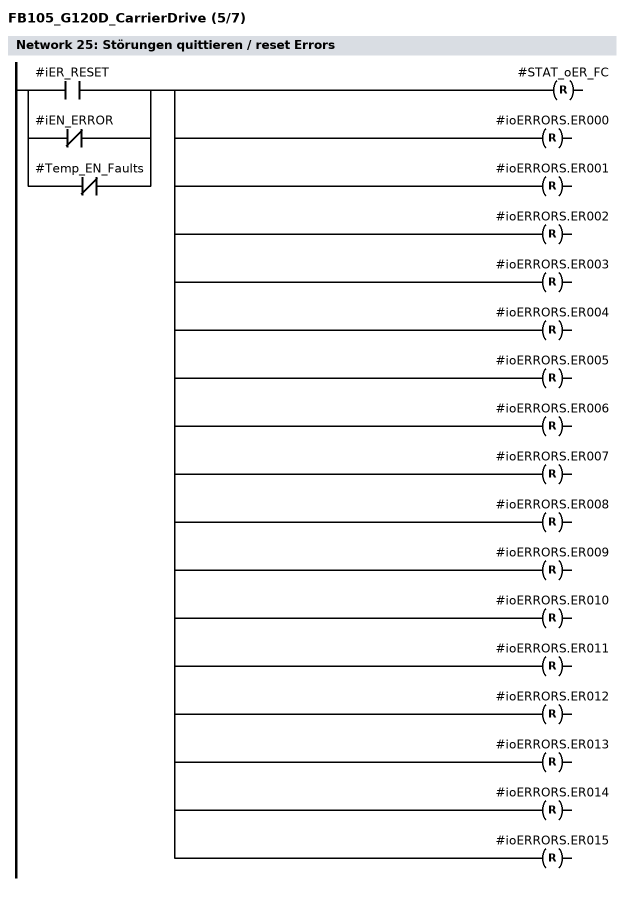
   RUNG wire#powerrail
      Contact( #iER_RESET )
      wire#w1
      R_Coil( #STAT_oER_FC )
   END_RUNG
   RUNG wire#powerrail
      I_Contact( #iEN_ERROR )
   END_RUNG wire#w1
   RUNG wire#powerrail
      I_Contact( #Temp_EN_Faults )
   END_RUNG wire#w1
   RUNG wire#w1
      R_Coil( #ioERRORS.ER000 )
   END_RUNG
   RUNG wire#w1
      R_Coil( #ioERRORS.ER001 )
   END_RUNG
   RUNG wire#w1
      R_Coil( #ioERRORS.ER002 )
   END_RUNG
   RUNG wire#w1
      R_Coil( #ioERRORS.ER003 )
   END_RUNG
   RUNG wire#w1
      R_Coil( #ioERRORS.ER004 )
   END_RUNG
   RUNG wire#w1
      R_Coil( #ioERRORS.ER005 )
   END_RUNG
   RUNG wire#w1
      R_Coil( #ioERRORS.ER006 )
   END_RUNG
   RUNG wire#w1
      R_Coil( #ioERRORS.ER007 )
   END_RUNG
   RUNG wire#w1
      R_Coil( #ioERRORS.ER008 )
   END_RUNG
   RUNG wire#w1
      R_Coil( #ioERRORS.ER009 )
   END_RUNG
   RUNG wire#w1
      R_Coil( #ioERRORS.ER010 )
   END_RUNG
   RUNG wire#w1
      R_Coil( #ioERRORS.ER011 )
   END_RUNG
   RUNG wire#w1
      R_Coil( #ioERRORS.ER012 )
   END_RUNG
   RUNG wire#w1
      R_Coil( #ioERRORS.ER013 )
   END_RUNG
   RUNG wire#w1
      R_Coil( #ioERRORS.ER014 )
   END_RUNG
   RUNG wire#w1
      R_Coil( #ioERRORS.ER015 )
   END_RUNG
   // the same network as SCL:
   IF #iER_RESET OR NOT #iEN_ERROR OR NOT #Temp_EN_Faults THEN
       #STAT_oER_FC := FALSE;
       #ioERRORS.ER000 := FALSE;
       #ioERRORS.ER001 := FALSE;
       #ioERRORS.ER002 := FALSE;
       #ioERRORS.ER003 := FALSE;
       #ioERRORS.ER004 := FALSE;
       #ioERRORS.ER005 := FALSE;
       #ioERRORS.ER006 := FALSE;
       #ioERRORS.ER007 := FALSE;
       #ioERRORS.ER008 := FALSE;
       #ioERRORS.ER009 := FALSE;
       #ioERRORS.ER010 := FALSE;
       #ioERRORS.ER011 := FALSE;
       #ioERRORS.ER012 := FALSE;
       #ioERRORS.ER013 := FALSE;
       #ioERRORS.ER014 := FALSE;
       #ioERRORS.ER015 := FALSE;
   END_IF;
END_REGION

REGION Network 26: Störungen / Errors
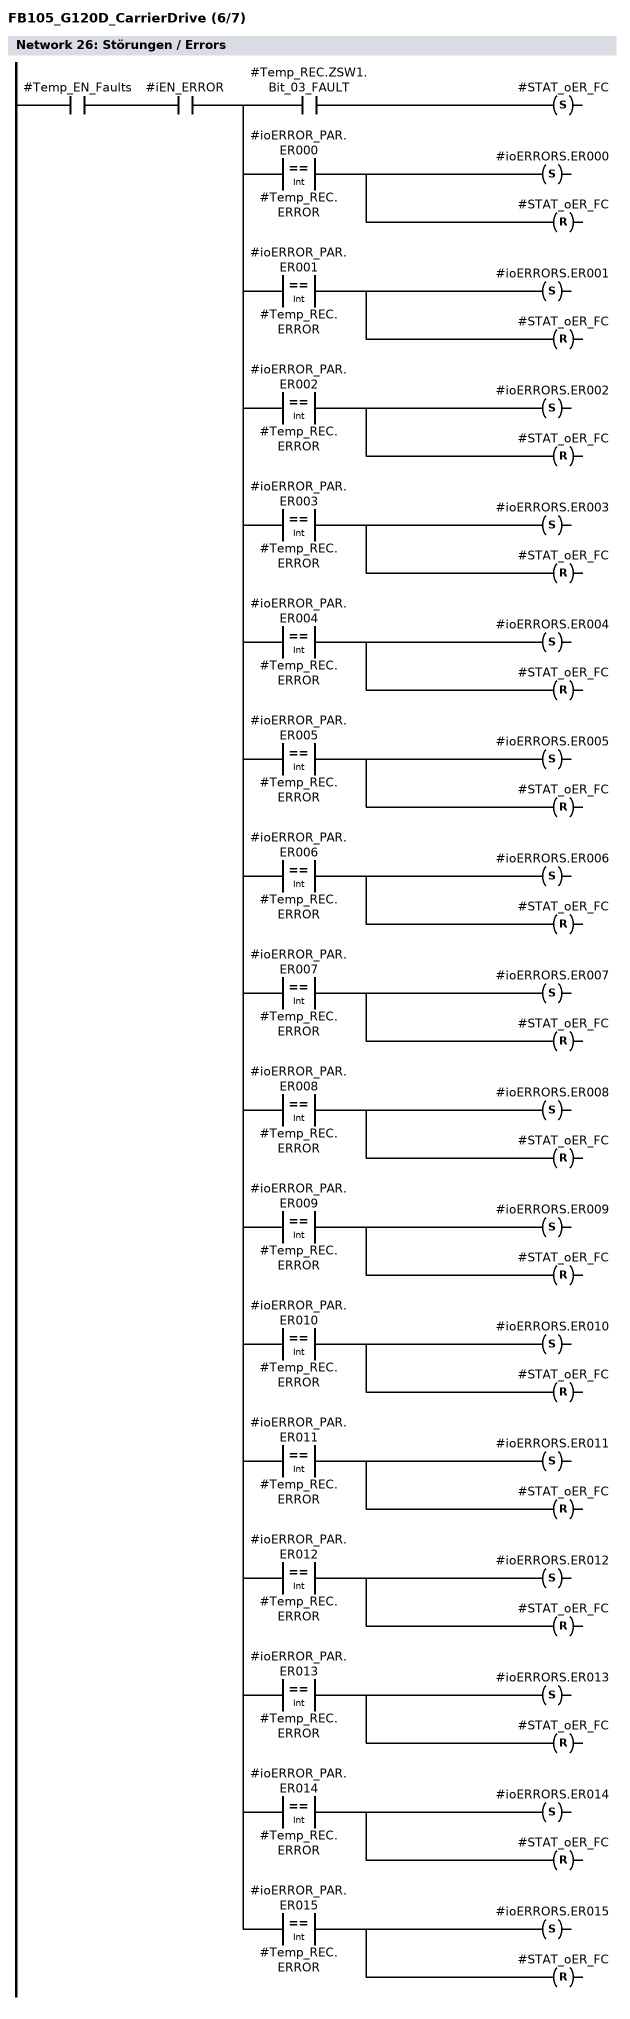
   RUNG wire#powerrail
      Contact( #Temp_EN_Faults )
      Contact( #iEN_ERROR )
      wire#w1
      Contact( #Temp_REC.ZSW1.Bit_03_FAULT )
      S_Coil( #STAT_oER_FC )
   END_RUNG
   RUNG wire#w1
      { S7_Templates := "SrcType := Int" } EQ_Contact(in1 := #ioERROR_PAR.ER000, in2 := #Temp_REC.ERROR)
      wire#w2
      S_Coil( #ioERRORS.ER000 )
   END_RUNG
   RUNG wire#w2
      R_Coil( #STAT_oER_FC )
   END_RUNG
   RUNG wire#w1
      { S7_Templates := "SrcType := Int" } EQ_Contact(in1 := #ioERROR_PAR.ER001, in2 := #Temp_REC.ERROR)
      wire#w3
      S_Coil( #ioERRORS.ER001 )
   END_RUNG
   RUNG wire#w3
      R_Coil( #STAT_oER_FC )
   END_RUNG
   RUNG wire#w1
      { S7_Templates := "SrcType := Int" } EQ_Contact(in1 := #ioERROR_PAR.ER002, in2 := #Temp_REC.ERROR)
      wire#w4
      S_Coil( #ioERRORS.ER002 )
   END_RUNG
   RUNG wire#w4
      R_Coil( #STAT_oER_FC )
   END_RUNG
   RUNG wire#w1
      { S7_Templates := "SrcType := Int" } EQ_Contact(in1 := #ioERROR_PAR.ER003, in2 := #Temp_REC.ERROR)
      wire#w5
      S_Coil( #ioERRORS.ER003 )
   END_RUNG
   RUNG wire#w5
      R_Coil( #STAT_oER_FC )
   END_RUNG
   RUNG wire#w1
      { S7_Templates := "SrcType := Int" } EQ_Contact(in1 := #ioERROR_PAR.ER004, in2 := #Temp_REC.ERROR)
      wire#w6
      S_Coil( #ioERRORS.ER004 )
   END_RUNG
   RUNG wire#w6
      R_Coil( #STAT_oER_FC )
   END_RUNG
   RUNG wire#w1
      { S7_Templates := "SrcType := Int" } EQ_Contact(in1 := #ioERROR_PAR.ER005, in2 := #Temp_REC.ERROR)
      wire#w7
      S_Coil( #ioERRORS.ER005 )
   END_RUNG
   RUNG wire#w7
      R_Coil( #STAT_oER_FC )
   END_RUNG
   RUNG wire#w1
      { S7_Templates := "SrcType := Int" } EQ_Contact(in1 := #ioERROR_PAR.ER006, in2 := #Temp_REC.ERROR)
      wire#w8
      S_Coil( #ioERRORS.ER006 )
   END_RUNG
   RUNG wire#w8
      R_Coil( #STAT_oER_FC )
   END_RUNG
   RUNG wire#w1
      { S7_Templates := "SrcType := Int" } EQ_Contact(in1 := #ioERROR_PAR.ER007, in2 := #Temp_REC.ERROR)
      wire#w9
      S_Coil( #ioERRORS.ER007 )
   END_RUNG
   RUNG wire#w9
      R_Coil( #STAT_oER_FC )
   END_RUNG
   RUNG wire#w1
      { S7_Templates := "SrcType := Int" } EQ_Contact(in1 := #ioERROR_PAR.ER008, in2 := #Temp_REC.ERROR)
      wire#w10
      S_Coil( #ioERRORS.ER008 )
   END_RUNG
   RUNG wire#w10
      R_Coil( #STAT_oER_FC )
   END_RUNG
   RUNG wire#w1
      { S7_Templates := "SrcType := Int" } EQ_Contact(in1 := #ioERROR_PAR.ER009, in2 := #Temp_REC.ERROR)
      wire#w11
      S_Coil( #ioERRORS.ER009 )
   END_RUNG
   RUNG wire#w11
      R_Coil( #STAT_oER_FC )
   END_RUNG
   RUNG wire#w1
      { S7_Templates := "SrcType := Int" } EQ_Contact(in1 := #ioERROR_PAR.ER010, in2 := #Temp_REC.ERROR)
      wire#w12
      S_Coil( #ioERRORS.ER010 )
   END_RUNG
   RUNG wire#w12
      R_Coil( #STAT_oER_FC )
   END_RUNG
   RUNG wire#w1
      { S7_Templates := "SrcType := Int" } EQ_Contact(in1 := #ioERROR_PAR.ER011, in2 := #Temp_REC.ERROR)
      wire#w13
      S_Coil( #ioERRORS.ER011 )
   END_RUNG
   RUNG wire#w13
      R_Coil( #STAT_oER_FC )
   END_RUNG
   RUNG wire#w1
      { S7_Templates := "SrcType := Int" } EQ_Contact(in1 := #ioERROR_PAR.ER012, in2 := #Temp_REC.ERROR)
      wire#w14
      S_Coil( #ioERRORS.ER012 )
   END_RUNG
   RUNG wire#w14
      R_Coil( #STAT_oER_FC )
   END_RUNG
   RUNG wire#w1
      { S7_Templates := "SrcType := Int" } EQ_Contact(in1 := #ioERROR_PAR.ER013, in2 := #Temp_REC.ERROR)
      wire#w15
      S_Coil( #ioERRORS.ER013 )
   END_RUNG
   RUNG wire#w15
      R_Coil( #STAT_oER_FC )
   END_RUNG
   RUNG wire#w1
      { S7_Templates := "SrcType := Int" } EQ_Contact(in1 := #ioERROR_PAR.ER014, in2 := #Temp_REC.ERROR)
      wire#w16
      S_Coil( #ioERRORS.ER014 )
   END_RUNG
   RUNG wire#w16
      R_Coil( #STAT_oER_FC )
   END_RUNG
   RUNG wire#w1
      { S7_Templates := "SrcType := Int" } EQ_Contact(in1 := #ioERROR_PAR.ER015, in2 := #Temp_REC.ERROR)
      wire#w17
      S_Coil( #ioERRORS.ER015 )
   END_RUNG
   RUNG wire#w17
      R_Coil( #STAT_oER_FC )
   END_RUNG
   // the same network as SCL:
   #_w1 := #Temp_EN_Faults AND #iEN_ERROR;
   IF #_w1 AND #Temp_REC.ZSW1.Bit_03_FAULT THEN #STAT_oER_FC := TRUE; END_IF;
   IF #_w1 AND (#ioERROR_PAR.ER000 = #Temp_REC.ERROR) THEN
       #ioERRORS.ER000 := TRUE;
       #STAT_oER_FC := FALSE;
   END_IF;
   IF #_w1 AND (#ioERROR_PAR.ER001 = #Temp_REC.ERROR) THEN
       #ioERRORS.ER001 := TRUE;
       #STAT_oER_FC := FALSE;
   END_IF;
   IF #_w1 AND (#ioERROR_PAR.ER002 = #Temp_REC.ERROR) THEN
       #ioERRORS.ER002 := TRUE;
       #STAT_oER_FC := FALSE;
   END_IF;
   IF #_w1 AND (#ioERROR_PAR.ER003 = #Temp_REC.ERROR) THEN
       #ioERRORS.ER003 := TRUE;
       #STAT_oER_FC := FALSE;
   END_IF;
   IF #_w1 AND (#ioERROR_PAR.ER004 = #Temp_REC.ERROR) THEN
       #ioERRORS.ER004 := TRUE;
       #STAT_oER_FC := FALSE;
   END_IF;
   IF #_w1 AND (#ioERROR_PAR.ER005 = #Temp_REC.ERROR) THEN
       #ioERRORS.ER005 := TRUE;
       #STAT_oER_FC := FALSE;
   END_IF;
   IF #_w1 AND (#ioERROR_PAR.ER006 = #Temp_REC.ERROR) THEN
       #ioERRORS.ER006 := TRUE;
       #STAT_oER_FC := FALSE;
   END_IF;
   IF #_w1 AND (#ioERROR_PAR.ER007 = #Temp_REC.ERROR) THEN
       #ioERRORS.ER007 := TRUE;
       #STAT_oER_FC := FALSE;
   END_IF;
   IF #_w1 AND (#ioERROR_PAR.ER008 = #Temp_REC.ERROR) THEN
       #ioERRORS.ER008 := TRUE;
       #STAT_oER_FC := FALSE;
   END_IF;
   IF #_w1 AND (#ioERROR_PAR.ER009 = #Temp_REC.ERROR) THEN
       #ioERRORS.ER009 := TRUE;
       #STAT_oER_FC := FALSE;
   END_IF;
   IF #_w1 AND (#ioERROR_PAR.ER010 = #Temp_REC.ERROR) THEN
       #ioERRORS.ER010 := TRUE;
       #STAT_oER_FC := FALSE;
   END_IF;
   IF #_w1 AND (#ioERROR_PAR.ER011 = #Temp_REC.ERROR) THEN
       #ioERRORS.ER011 := TRUE;
       #STAT_oER_FC := FALSE;
   END_IF;
   IF #_w1 AND (#ioERROR_PAR.ER012 = #Temp_REC.ERROR) THEN
       #ioERRORS.ER012 := TRUE;
       #STAT_oER_FC := FALSE;
   END_IF;
   IF #_w1 AND (#ioERROR_PAR.ER013 = #Temp_REC.ERROR) THEN
       #ioERRORS.ER013 := TRUE;
       #STAT_oER_FC := FALSE;
   END_IF;
   IF #_w1 AND (#ioERROR_PAR.ER014 = #Temp_REC.ERROR) THEN
       #ioERRORS.ER014 := TRUE;
       #STAT_oER_FC := FALSE;
   END_IF;
   IF #_w1 AND (#ioERROR_PAR.ER015 = #Temp_REC.ERROR) THEN
       #ioERRORS.ER015 := TRUE;
       #STAT_oER_FC := FALSE;
   END_IF;
END_REGION

REGION Network 27: OUT: Störung FU allgemein
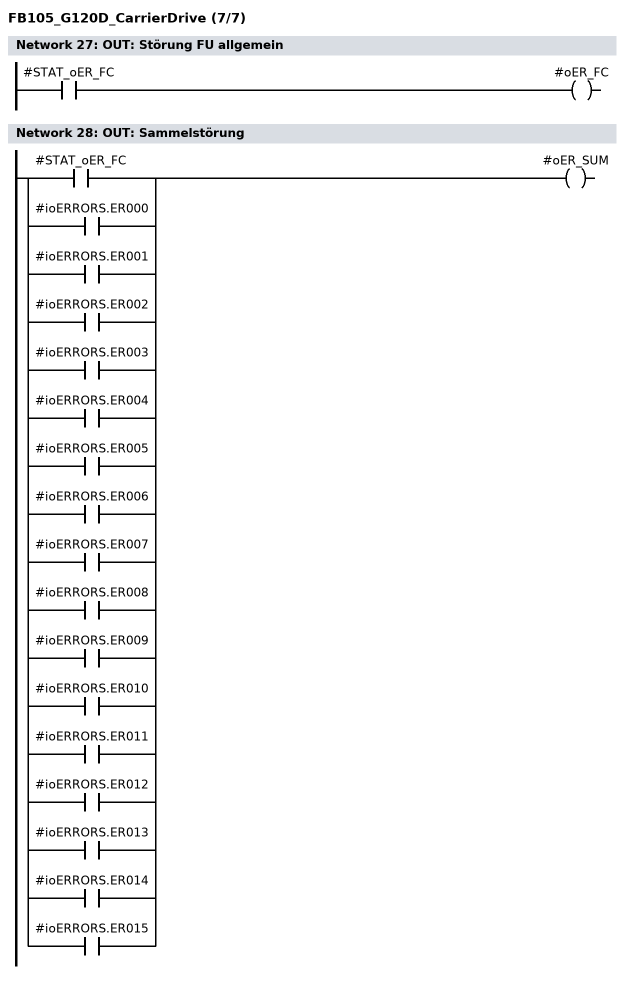
   RUNG wire#powerrail
      Contact( #STAT_oER_FC )
      Coil( #oER_FC )
   END_RUNG
   // the same network as SCL:
   #oER_FC := #STAT_oER_FC;
END_REGION

REGION Network 28: OUT: Sammelstörung
   RUNG wire#powerrail
      Contact( #STAT_oER_FC )
      wire#w1
      Coil( #oER_SUM )
   END_RUNG
   RUNG wire#powerrail
      Contact( #ioERRORS.ER000 )
   END_RUNG wire#w1
   RUNG wire#powerrail
      Contact( #ioERRORS.ER001 )
   END_RUNG wire#w1
   RUNG wire#powerrail
      Contact( #ioERRORS.ER002 )
   END_RUNG wire#w1
   RUNG wire#powerrail
      Contact( #ioERRORS.ER003 )
   END_RUNG wire#w1
   RUNG wire#powerrail
      Contact( #ioERRORS.ER004 )
   END_RUNG wire#w1
   RUNG wire#powerrail
      Contact( #ioERRORS.ER005 )
   END_RUNG wire#w1
   RUNG wire#powerrail
      Contact( #ioERRORS.ER006 )
   END_RUNG wire#w1
   RUNG wire#powerrail
      Contact( #ioERRORS.ER007 )
   END_RUNG wire#w1
   RUNG wire#powerrail
      Contact( #ioERRORS.ER008 )
   END_RUNG wire#w1
   RUNG wire#powerrail
      Contact( #ioERRORS.ER009 )
   END_RUNG wire#w1
   RUNG wire#powerrail
      Contact( #ioERRORS.ER010 )
   END_RUNG wire#w1
   RUNG wire#powerrail
      Contact( #ioERRORS.ER011 )
   END_RUNG wire#w1
   RUNG wire#powerrail
      Contact( #ioERRORS.ER012 )
   END_RUNG wire#w1
   RUNG wire#powerrail
      Contact( #ioERRORS.ER013 )
   END_RUNG wire#w1
   RUNG wire#powerrail
      Contact( #ioERRORS.ER014 )
   END_RUNG wire#w1
   RUNG wire#powerrail
      Contact( #ioERRORS.ER015 )
   END_RUNG wire#w1
   // the same network as SCL:
   #oER_SUM := #STAT_oER_FC OR #ioERRORS.ER000 OR #ioERRORS.ER001 OR #ioERRORS.ER002 OR #ioERRORS.ER003 OR #ioERRORS.ER004 OR #ioERRORS.ER005 OR #ioERRORS.ER006 OR #ioERRORS.ER007 OR #ioERRORS.ER008 OR #ioERRORS.ER009 OR #ioERRORS.ER010 OR #ioERRORS.ER011 OR #ioERRORS.ER012 OR #ioERRORS.ER013 OR #ioERRORS.ER014 OR #ioERRORS.ER015;
END_REGION

REGION Network 29: ENDE / END
   // ################################ ENDE ############################### / ###################################### END #####################################
END_REGION
END_FUNCTION_BLOCK

FUNCTION_BLOCK "FB1110_Red_Green_LED"   // FB1110, LAD
{ S7_Optimized_Access := 'TRUE' }
VERSION : 0.1
   VAR_INPUT
      Red : Bool;
      Green : Bool;
   END_VAR
   VAR
      instWRREC : WRREC;
      statWRREC_LEDByte : Byte;
   END_VAR
BEGIN

REGION Network 1: Red LED
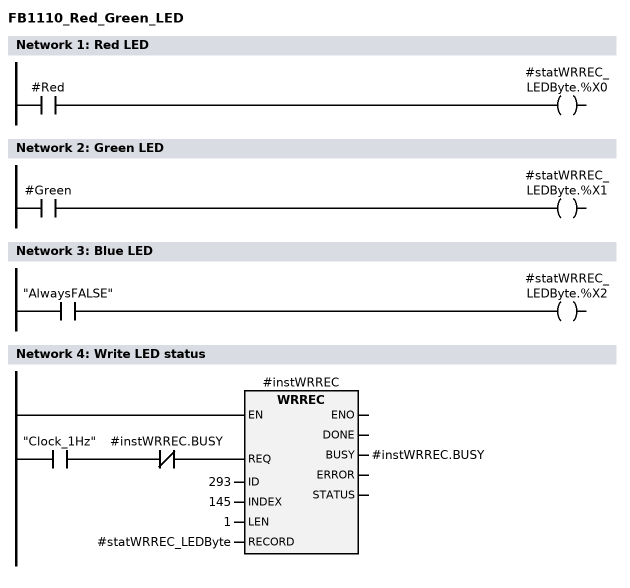
   RUNG wire#powerrail
      Contact( #Red )
      Coil( #statWRREC_LEDByte.%X0 )
   END_RUNG
   // the same network as SCL:
   #statWRREC_LEDByte.%X0 := #Red;
END_REGION

REGION Network 2: Green LED
   RUNG wire#powerrail
      Contact( #Green )
      Coil( #statWRREC_LEDByte.%X1 )
   END_RUNG
   // the same network as SCL:
   #statWRREC_LEDByte.%X1 := #Green;
END_REGION

REGION Network 3: Blue LED
   RUNG wire#powerrail
      Contact( "AlwaysFALSE" )
      Coil( #statWRREC_LEDByte.%X2 )
   END_RUNG
   // the same network as SCL:
   #statWRREC_LEDByte.%X2 := "AlwaysFALSE";
END_REGION

REGION Network 4: Write LED status
   #instWRREC(REQ := "Clock_1Hz" AND NOT #instWRREC.BUSY,   // WRREC
              ID := 293,
              INDEX := 145,
              LEN := 1,
              RECORD := #statWRREC_LEDByte,
              BUSY => #instWRREC.BUSY);
END_REGION

REGION Network 5: End
END_REGION
END_FUNCTION_BLOCK

// folder: 03_FB'S/DIAGNOSTICS

FUNCTION_BLOCK "FB1000_Default_SupervisionFB"   // FB1000, ProDiag
{ S7_Optimized_Access := 'TRUE' }
   VAR
      State : SV_FB_State;
   END_VAR
   VAR_TEMP
      t_TempSvStateUDT : SV_State;
      t_TempAlarmInstance : <type 200004f>;
      t_TempAsocValue1 : Variant;
      t_TempAsocValue2 : Variant;
      t_TempAsocValue3 : Variant;
   END_VAR
BEGIN
END_FUNCTION_BLOCK

FUNCTION_BLOCK "FB1001_EMS_BreakerStatus"   // FB1001, LAD
TITLE = Monitoring Fuse
{ S7_Optimized_Access := 'TRUE' }
AUTHOR : Siemens
FAMILY : LSimoveC
VERSION : 1.0
// © 2018 Siemens AG 
// SIMOVE Carrier Control
   VAR_INPUT
      Diag : Variant;   // Diagnosis signal of the selectivity module
   END_VAR
   VAR_OUTPUT
      Channel1 : Bool;   // Channel 1 active
      Channel2 : Bool;   // Channel 2 active
      Channel3 : Bool;   // Channel 3 active
      Channel4 : Bool;   // Channel 4 active
      CollectiveError : Bool;   // Collective error of the selectivity module
   END_VAR
   VAR
      instDiagBreaker : "FB1002_LSimoveC_DiagBreaker";
      instTimeout : TON_TIME;
      statError : Bool;
   END_VAR
   VAR_TEMP
      tempDone : Bool;
      tempBusy : Bool;
      tempChannelState : Byte;
      tempStatus : Word;
      tempDiag : Bool;
      tempInt : Int;
      tempModuleOK : Bool;
      tempHW : Hw_Any;
      tempDiagInfo : DIS;
      tempUInt : UInt;
      tempTimeout : Bool;
   END_VAR
BEGIN

REGION Network 1: Change journal
   // =============================================================================
   // Siemens AG
   // (c)Copyright 2018 Alle Rechte vorbehalten
   // -----------------------------------------------------------------------------
   // Bibliothek: LSimoveC
   // Funktion: Der FB wertet den Status-Ausgang eines SITOP-Selektivitätsmoduls aus. Der Status-Ausgang liefert ein Signal, das den Zustand der Verbaucherkreise seriell codiert. Der Baustein decodiert das Signal und stellt den Status der Verbraucherkreise als Einzelsignale zur Verfügung.
   // -----------------------------------------------------------------------------
   // Änderungsjournal:
   // V1.0  01.02.2018  Neuerstellung
   // =============================================================================
END_REGION

REGION Network 2: Determine block error
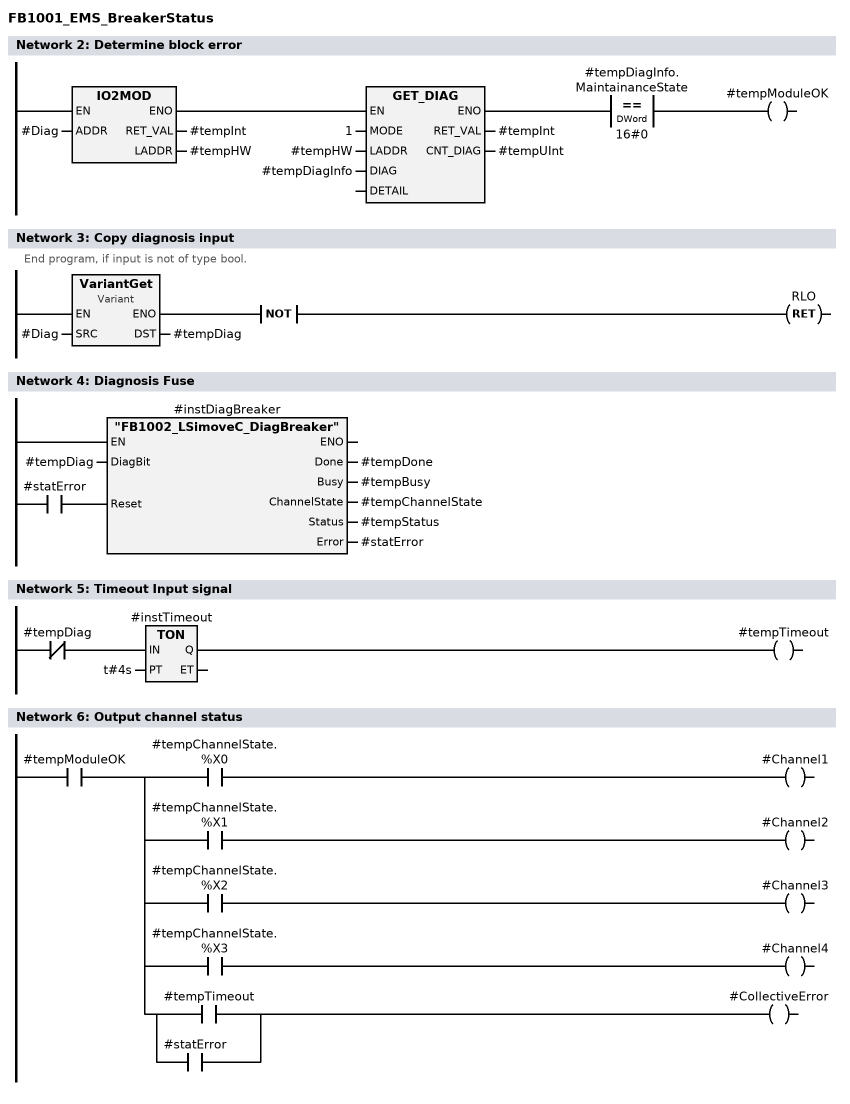
   // ENO of a box is taken as its EN; it also drops when the box reports an error
   #tempInt := IO2MOD(ADDR := #Diag, LADDR => #tempHW);
   #tempInt := GET_DIAG(MODE := 1, LADDR := #tempHW, DIAG := #tempDiagInfo, CNT_DIAG => #tempUInt);
   #tempModuleOK := #tempDiagInfo.MaintainanceState = 16#0;
END_REGION

REGION Network 3: Copy diagnosis input
   // End program, if input is not of type bool.
   // no SCL statement known for VariantGet: written as a call
   // ENO of a box is taken as its EN; it also drops when the box reports an error
   VariantGet(src := #Diag, dst => #tempDiag);
   IF NOT TRUE THEN
       ENO := TRUE;
       RETURN;
   END_IF;
END_REGION

REGION Network 4: Diagnosis Fuse
   RUNG wire#powerrail
      #instDiagBreaker(Reset := wire#w1, DiagBit := #tempDiag, Done => #tempDone, Busy => #tempBusy, ChannelState => #tempChannelState, Status => #tempStatus, Error => #statError)
   END_RUNG
   RUNG wire#powerrail
      Contact( #statError )
   END_RUNG wire#w1
   // the same network as SCL:
   #instDiagBreaker(DiagBit := #tempDiag,   // "FB1002_LSimoveC_DiagBreaker"
                    Reset := #statError,
                    Done => #tempDone,
                    Busy => #tempBusy,
                    ChannelState => #tempChannelState,
                    Status => #tempStatus,
                    Error => #statError);
END_REGION

REGION Network 5: Timeout Input signal
   #instTimeout(IN := NOT #tempDiag, PT := t#4s);   // TON
   #tempTimeout := #instTimeout.Q;
END_REGION

REGION Network 6: Output channel status
   RUNG wire#powerrail
      Contact( #tempModuleOK )
      wire#w1
      Contact( #tempChannelState.%X0 )
      Coil( #Channel1 )
   END_RUNG
   RUNG wire#w1
      Contact( #tempChannelState.%X1 )
      Coil( #Channel2 )
   END_RUNG
   RUNG wire#w1
      Contact( #tempChannelState.%X2 )
      Coil( #Channel3 )
   END_RUNG
   RUNG wire#w1
      Contact( #tempChannelState.%X3 )
      Coil( #Channel4 )
   END_RUNG
   RUNG wire#w1
      Contact( #tempTimeout )
      wire#w2
      Coil( #CollectiveError )
   END_RUNG
   RUNG wire#w1
      Contact( #statError )
   END_RUNG wire#w2
   // the same network as SCL:
   #Channel1 := #tempModuleOK AND #tempChannelState.%X0;
   #Channel2 := #tempModuleOK AND #tempChannelState.%X1;
   #Channel3 := #tempModuleOK AND #tempChannelState.%X2;
   #Channel4 := #tempModuleOK AND #tempChannelState.%X3;
   #CollectiveError := #tempModuleOK AND (#tempTimeout OR #statError);
END_REGION
END_FUNCTION_BLOCK

FUNCTION_BLOCK "FB1002_LSimoveC_DiagBreaker"   // FB1002, SCL
TITLE = DiagnoseSicherung
{ S7_Optimized_Access := 'FALSE' }
AUTHOR : Siemens
FAMILY : LSimoveC
VERSION : 2.3
// © 2018 Siemens AG 
// SIMOVE Carrier Control
   VAR_INPUT
      DiagBit : Bool;   // Input through which the signal of the status output of the selectivity module is read
      Reset : Bool;   // A positive edge triggers a reset. All parameters are reset.
   END_VAR
   VAR_OUTPUT
      Done : Bool;   // Done = 1: A telegram was evaluated completely and without errors. Done = 0: telegram evaluation is running or no signal is detected at the input "impulse".
      Busy : Bool;   // Busy = 1: Function module "LSitop_PseDiag" is active. Busy = 0: if done=1, a telegram was evaluated completely and without error.
      ChannelState : Byte;   // State of the outputs 1 to 4.
      Status : Word;   // Status display: if error=1, the error number for one cycle is displayed at the output "status". if error=0, the value 16 # 0000 is displayed at the output "status".
      Error : Bool;   // Error=1: an error has occured during the execution of the routine. The value error=1 is set for one cycle. if error=0: no error.
   END_VAR
   VAR
      statImpulseOld : Bool;
      statResetOld : Bool;
      statTimeSaver : Struct
         TimeTckRisingEdge : Time;
         TimeTckFallingEdge : Time;
         RisingEdgeDetected : Bool;
         FallingEdgeDetected : Bool;
         stateEdge : Int := 0;
      END_STRUCT;
      statDeltaTimeImpulse : Time;
      statDeltaTimePause : Time;
      statStartImpulseDetected : Bool;
      statImpulseDetected : Bool;
      statChannelState : Byte;
      statTimePauseSave0 : Time;
      statTimePauseSave1 : Time;
      statTimePauseSave2 : Time;
      statTimePauseSave3 : Time;
      statTimePauseSave4 : Time;
      statTimeImpulseSave0 : Time;
      statTimeImpulseSave1 : Time;
      statTimeImpulseSave2 : Time;
      statTimeImpulseSave3 : Time;
      statTimeImpulseSave4 : Time;
      statFrameImulseDetected : Bool;
      statNumberOfImpulses : Int;
      statChannelActive1 : Bool;
      statChannelActive2 : Bool;
      statChannelActive3 : Bool;
      statChannelActive4 : Bool;
      statCountChannelPos : Int;
      statCurrentPos1 : Int;
      statCurrentPos2 : Int;
      statCurrentPos3 : Int;
      statCurrentPos4 : Int;
      statTimeToImpulse : Time;
      statTimePause : Time;
      statTimeImpulse : Time;
      statTimeFrame : Time;
      statFrameOk : Bool;
      statCycleTimeNok : Bool;
      statSysTime : Time;
      statSysTimeOld : Time;
      statDeltaSysTime : Time;
      instSysTimer : TON_TIME;
      statSysTimerStart : Bool;
      statSysTimerStop : Bool;
      statStatus : Word;
      statIndex : Int;
      statSysTimerRun : Time;
      instWatchDogTimerRising : TON_TIME;
      statWatchDogTimerRisingStart : Bool;
      statWatchDogTimerRisingStop : Bool;
      statWatchDogTimerRisingRun : Time;
      statResetRequest : Bool;
      instWatchDogTimerFalling : TON_TIME;
      statWatchDogTimerFallingStart : Bool;
      statWatchDogTimerFallingStop : Bool;
      statWatchDogTimerFallingRun : Time;
   END_VAR
   VAR_TEMP
      tempLatchTime : Time;
   END_VAR
   VAR CONSTANT
      STATE_IDLE : Int := 0;
      STATE_EVALUATION : Int := 1;
      STATE_ERROR : Int := 2;
      TIME_FRAME_MAX : Time := T#2850ms;
      TIME_FRAME_MIN : Time := T#2650ms;
      TIME_STARTIMPULSE_MAX : Time := T#600ms;
      TIME_STARTIMPULSE_MIN : Time := T#400ms;
      TIME_IMPULSE_MIN : Time := T#150ms;
      TIME_IMPULSE_MAX : Time := T#350ms;
      TIME_PAUSE1_MIN : Time := T#150ms;
      TIME_PAUSE1_MAX : Time := T#350ms;
      TIME_PAUSE2_MIN : Time := T#650ms;
      TIME_PAUSE2_MAX : Time := T#850ms;
      TIME_PAUSE3_MIN : Time := T#1150ms;
      TIME_PAUSE3_MAX : Time := T#1350ms;
      TIME_PAUSE4_MIN : Time := T#1650ms;
      TIME_PAUSE4_MAX : Time := T#1850ms;
      TIME_PAUSE_FRAME_MAX : Time := T#2350ms;
      TIME_PAUSE_FRAME_MIN : Time := T#2150ms;
      TIME_CONST_0 : Time := T#0ms;
      TIME_CONST_102 : Time := T#102ms;
      CONST_STATE_RISING_EDGE : Int := 15;
      CONST_STATE_FALLING_EDGE : Int := 16;
      CONST_WORD_0 : Word := 16#0000;
      CONST_BYTE_0 : Byte := 16#00;
      CONST_INT_0 : Int := 0;
      CONST_CHANNEL_POS4 : Int := 4;
      CONST_CHANNEL_POS1 : Int := 1;
      CONST_CHANNEL_POS2 : Int := 2;
      CONST_CHANNEL_POS3 : Int := 3;
      CONST_WATCHDOG_TIMER : Time := T#6s;
      CONST_CYCLETIME_TIMER : Time := t#4s;
      CONST_ERROR_CYCLETIME_TIMER : Word := 16#8001;
      CONST_ERROR_WATCHDOG_TIMER : Word := 16#8002;
   END_VAR
BEGIN
   //=============================================================================
   //SIEMENES AG
   //(c)Copyright 2017 All Rights Reserved
   //-----------------------------------------------------------------------------
   //Library:       LSitop
   //Tested with:   (S7-1500)
   //Engineering:    TIA Portal V14
   //Restrictions:   call in cyclic main OB
   //Requirements:
   //Functionality: evaluates the signal of status output (S) of SITOP PSE200U 
   //               ....
   //
   //-----------------------------------------------------------------------------
   //Change log table:
   //Version  Date       Expert in charge Changes applied
   //02.03.01 24.05.2017 (DF CS SD CCC OS) Third released version
   //=============================================================================

   // Calculate cycle time
   #statSysTime:=TIME_TCK();
   #statDeltaSysTime := #statSysTime - #statSysTimeOld;

   IF (#statDeltaSysTime < t#0ms)
   THEN
       #statDeltaSysTime := #statDeltaSysTime + T#2147483647ms;

       IF (#statDeltaSysTime < #TIME_CONST_0)
       THEN
           #statCycleTimeNok := true;
           #statSysTimeOld := #statSysTime;
           RETURN;
       ELSE
           #statCycleTimeNok := false;
       END_IF;

   ELSIF (#statDeltaSysTime >= #TIME_CONST_102)
   THEN
       #statCycleTimeNok := true;
       #statSysTimerStart := true;
   ELSE
       #statCycleTimeNok := false;
       #statSysTimerStart := false;
   END_IF;

   //Rising edge at reset input

   IF ((#Reset = true)
       AND (#statResetOld = false))
   THEN
       #statSysTimerStart := false;
       #statWatchDogTimerRisingStart := false;
       #statWatchDogTimerFallingStart := false;
       #statResetRequest := true;
       #statIndex := #STATE_IDLE;
   END_IF;

   //Rising edge at impulse input
   IF ((#DiagBit = True)
       AND (#statImpulseOld = False))
   THEN
       #tempLatchTime := TIME_TCK();
       #statTimeSaver.RisingEdgeDetected := true;
       #statTimeSaver.stateEdge := #CONST_STATE_RISING_EDGE;
       #statTimeSaver.TimeTckRisingEdge := #tempLatchTime;
       #statWatchDogTimerRisingStart := true;
       #statWatchDogTimerFallingStart := false;

       IF (#Busy = false)
       THEN
           #Busy := true;
           #Done := false;
           #Error := false;
           #Status := #CONST_WORD_0;
       END_IF;

       IF ((#statCycleTimeNok = false)
           AND (#statResetRequest = false))
       THEN
           #statIndex := #STATE_EVALUATION;
       END_IF;

   END_IF;

   //Falling edge at impulse input
   IF ((#DiagBit = False)
       AND (#statImpulseOld = True))
   THEN
       #tempLatchTime := TIME_TCK();
       #statTimeSaver.FallingEdgeDetected := true;
       #statTimeSaver.stateEdge := #CONST_STATE_FALLING_EDGE;
       #statTimeSaver.TimeTckFallingEdge := #tempLatchTime;

       #statWatchDogTimerFallingStart := true;
       #statWatchDogTimerRisingStart := false;

       IF ((#statCycleTimeNok = FALSE)
           AND (#statResetRequest = false))
       THEN
           #statIndex := #STATE_EVALUATION;
       END_IF;

   END_IF;

   IF ((#statTimeSaver.FallingEdgeDetected = false)
       AND (#statTimeSaver.RisingEdgeDetected = FALSE))
   THEN
       #statWatchDogTimerRisingStart := true;
       #statWatchDogTimerFallingStart := true;
   END_IF;

   CASE #statIndex OF
       #STATE_IDLE:  // IDLE_STATE
           #Done := false;
           #Error := false;
           #Busy := false;
           #Status := #CONST_WORD_0;
           #statStatus := #CONST_WORD_0;
           #ChannelState := #CONST_BYTE_0;
           #statChannelState := #CONST_BYTE_0;
           #statFrameOk := false;
           #statCycleTimeNok := false;
           #statStartImpulseDetected := false;
           #statFrameImulseDetected := false;
           #statResetRequest := false;
           #statTimeSaver.FallingEdgeDetected := false;
           #statTimeSaver.RisingEdgeDetected := false;

       #STATE_EVALUATION:  //State: impulse detection

           //Delta time calculation
           IF ((#statTimeSaver.RisingEdgeDetected = True)
               AND (#statTimeSaver.FallingEdgeDetected = True))
           THEN

               IF (#statTimeSaver.stateEdge = #CONST_STATE_RISING_EDGE) //pos. edge, evaluate delta pause
               THEN
                   #statDeltaTimePause := #statTimeSaver.TimeTckRisingEdge - #statTimeSaver.TimeTckFallingEdge;

                   IF (#statDeltaTimePause < #TIME_CONST_0)
                   THEN
                       #statDeltaTimePause := #statDeltaTimePause + T#2147483647ms;

                       IF (#statDeltaTimePause < #TIME_CONST_0)
                       THEN
                           #statIndex := #STATE_IDLE;
                           #statTimeSaver.FallingEdgeDetected := false;
                           RETURN;
                       END_IF;

                   ELSIF (#statDeltaTimePause > #TIME_FRAME_MAX)
                   THEN
                       #statIndex := #STATE_IDLE;
                       #statTimeSaver.FallingEdgeDetected := false;
                       RETURN;
                   END_IF;
                   #statTimeSaver.FallingEdgeDetected := false;
               END_IF;

               IF (#statTimeSaver.stateEdge = #CONST_STATE_FALLING_EDGE) // neg. edge, evaluate delta impulse
               THEN
                   #statImpulseDetected := true;
                   #statDeltaTimeImpulse := #statTimeSaver.TimeTckFallingEdge - #statTimeSaver.TimeTckRisingEdge;

                   IF (#statDeltaTimeImpulse < #TIME_CONST_0)
                   THEN
                       #statDeltaTimeImpulse := #statDeltaTimeImpulse + T#2147483647ms;

                       IF (#statDeltaTimeImpulse < #TIME_CONST_0)
                       THEN
                           #statIndex := #STATE_IDLE;
                           #statTimeSaver.RisingEdgeDetected := false;
                           RETURN;
                       END_IF;

                   ELSIF (#statDeltaTimeImpulse > #TIME_FRAME_MAX)
                   THEN
                       #statIndex := #STATE_IDLE;
                       #statTimeSaver.RisingEdgeDetected := false;
                       RETURN;
                   END_IF;
                   #statTimeSaver.RisingEdgeDetected := false;
               END_IF;
           END_IF;

           //Start bit detection
           IF ((#statDeltaTimeImpulse >= #TIME_STARTIMPULSE_MIN)
               AND (#statDeltaTimeImpulse <= #TIME_STARTIMPULSE_MAX))
               AND (#statImpulseDetected = True)
           THEN
               #statImpulseDetected := False;
               #statNumberOfImpulses := #CONST_INT_0;
               #statCountChannelPos := #CONST_INT_0;

               IF (#statCurrentPos1 = #CONST_INT_0)
               THEN
                   #statTimeImpulseSave1 := #TIME_CONST_0;
                   #statTimePauseSave1 := #TIME_CONST_0;
               END_IF;

               IF (#statCurrentPos2 = #CONST_INT_0)
               THEN
                   #statTimeImpulseSave2 := #TIME_CONST_0;
                   #statTimePauseSave2 := #TIME_CONST_0;
               END_IF;

               IF (#statCurrentPos3 = #CONST_INT_0)
               THEN
                   #statTimeImpulseSave3 := #TIME_CONST_0;
                   #statTimePauseSave3 := #TIME_CONST_0;
               END_IF;

               IF (#statCurrentPos4 = #CONST_INT_0)
               THEN
                   #statTimeImpulseSave4 := #TIME_CONST_0;
                   #statTimePauseSave4 := #TIME_CONST_0;
               END_IF;

               #statTimePauseSave0 := #statDeltaTimePause;
               #statTimeImpulseSave0 := #statDeltaTimeImpulse;

               // get time in sum of imulses
               #statTimeImpulse := #statTimeImpulseSave0 + #statTimeImpulseSave1 + #statTimeImpulseSave2 + #statTimeImpulseSave3 + #statTimeImpulseSave4;

               //get time in sum of pauses
               #statTimePause := #statTimePauseSave0 + #statTimePauseSave1 + #statTimePauseSave2 + #statTimePauseSave3 + #statTimePauseSave4;

               // get length of frame
               #statTimeFrame := #statTimeImpulse + #statTimePause;

               IF ((#statTimeFrame >= #TIME_FRAME_MIN)
                   AND (#statTimeFrame <= #TIME_FRAME_MAX)
                   AND (#statTimeToImpulse <= #TIME_FRAME_MAX))
               THEN
                   #statFrameOk := true;
               END_IF;

               IF ((#statFrameOk = TRUE)
                   AND (#statCycleTimeNok = FALSE))
               THEN
                   // take over data
                   #Done := true;
                   #Busy := false;
                   #statFrameOk := false;

                   IF (#statChannelActive1 = true)
                   THEN
                       #statChannelState.%X0 := false;
                   ELSE
                       #statChannelState.%X0 := true;
                   END_IF;

                   IF (#statChannelActive2 = true)
                   THEN
                       #statChannelState.%X1 := false;
                   ELSE
                       #statChannelState.%X1 := true;
                   END_IF;

                   IF (#statChannelActive3 = true)
                   THEN
                       #statChannelState.%X2 := false;
                   ELSE
                       #statChannelState.%X2 := true;
                   END_IF;

                   IF (#statChannelActive4 = true)
                   THEN
                       #statChannelState.%X3 := false;
                   ELSE
                       #statChannelState.%X3 := true;
                   END_IF;

                   #ChannelState := #statChannelState;
               END_IF;


               // channel 4 ok
               IF ((#statDeltaTimePause >= #TIME_PAUSE1_MIN)
                   AND (#statDeltaTimePause <= #TIME_PAUSE1_MAX))
               THEN
                   #statChannelActive4 := true;
                   // channel 4 ok not ok
               ELSIF ((#statDeltaTimePause >= #TIME_PAUSE2_MIN)
                   AND (#statDeltaTimePause <= #TIME_PAUSE2_MAX))
               THEN
                   #statChannelActive4 := false;
                   // channel 3 and 4 not ok    
               ELSIF ((#statDeltaTimePause >= #TIME_PAUSE3_MIN)
                   AND (#statDeltaTimePause <= #TIME_PAUSE3_MAX))
               THEN
                   #statChannelActive3 := false;
                   #statChannelActive4 := false;
                   // channel 2, 3, 4 not ok
               ELSIF ((#statDeltaTimePause >= #TIME_PAUSE4_MIN)
                   AND (#statDeltaTimePause <= #TIME_PAUSE4_MAX))
               THEN
                   #statChannelActive2 := false;
                   #statChannelActive3 := false;
                   #statChannelActive4 := false;
                   // channel 1, 2, 3, 4 not ok
               ELSIF ((#statDeltaTimePause >= #TIME_PAUSE_FRAME_MIN)
                   AND (#statDeltaTimePause <= #TIME_PAUSE_FRAME_MAX))
               THEN
                   #statChannelActive1 := false;
                   #statChannelActive2 := false;
                   #statChannelActive3 := false;
                   #statChannelActive4 := false;
               END_IF;

               #statCountChannelPos := #CONST_CHANNEL_POS4;

               #statCurrentPos1 := #CONST_INT_0;
               #statCurrentPos2 := #CONST_INT_0;
               #statCurrentPos3 := #CONST_INT_0;
               #statCurrentPos4 := #CONST_INT_0;

           // Imulse bit detection
           ELSIF ((#statDeltaTimeImpulse >= #TIME_IMPULSE_MIN)
               AND (#statDeltaTimeImpulse <= #TIME_IMPULSE_MAX))
               AND (#statImpulseDetected = True)
           THEN
               #statImpulseDetected := False;
               #statFrameImulseDetected := true;
           END_IF;

           //Channel detection
           IF #statFrameImulseDetected = TRUE
           THEN
               #statFrameImulseDetected := FALSE;

               IF (#statCountChannelPos = #CONST_CHANNEL_POS4)
               THEN
                   #statCurrentPos1 := #statCountChannelPos;
                   #statTimeImpulseSave1 := #statDeltaTimeImpulse;
                   #statTimePauseSave1 := #statDeltaTimePause;
                   #statTimeToImpulse := #TIME_CONST_0;
                   #statTimeToImpulse := #statTimeToImpulse + #statDeltaTimeImpulse + #statDeltaTimePause;

                   //channel 1 ok
                   IF ((#statDeltaTimePause >= #TIME_PAUSE1_MIN)
                       AND (#statDeltaTimePause <= #TIME_PAUSE1_MAX))
                   THEN
                       #statChannelActive1 := true;
                       #statCountChannelPos := #CONST_CHANNEL_POS1; // Pos 1 detected
                   END_IF;

                   // channel 1 not ok
                   IF ((#statDeltaTimePause >= #TIME_PAUSE2_MIN)
                       AND (#statDeltaTimePause <= #TIME_PAUSE2_MAX))
                   THEN
                       #statChannelActive1 := false;
                       #statChannelActive2 := true;
                       #statCountChannelPos := #CONST_CHANNEL_POS2; // go to next Pos 2
                   END_IF;

                   // channel 1 and 2 not ok
                   IF ((#statDeltaTimePause >= #TIME_PAUSE3_MIN)
                       AND (#statDeltaTimePause <= #TIME_PAUSE3_MAX))
                   THEN
                       #statChannelActive1 := false;
                       #statChannelActive2 := false;
                       #statChannelActive3 := true;
                       #statCountChannelPos := #CONST_CHANNEL_POS2; // go to next Pos 2
                   END_IF;

                   // channel 1, 2 and 3 not ok
                   IF ((#statDeltaTimePause >= #TIME_PAUSE4_MIN)
                       AND (#statDeltaTimePause <= #TIME_PAUSE4_MAX))
                   THEN
                       #statChannelActive1 := false;
                       #statChannelActive2 := false;
                       #statChannelActive3 := FALSE;
                       #statChannelActive4 := true;
                       #statCountChannelPos := #CONST_INT_0;
                   END_IF;

               ELSIF (#statCountChannelPos = #CONST_CHANNEL_POS1)
               THEN
                   #statCurrentPos2 := #statCountChannelPos;
                   #statTimeImpulseSave2 := #statDeltaTimeImpulse;
                   #statTimePauseSave2 := #statDeltaTimePause;
                   #statTimeToImpulse := #statTimeToImpulse + #statDeltaTimeImpulse + #statDeltaTimePause;

                   IF ((#statDeltaTimePause >= #TIME_PAUSE1_MIN)
                       AND (#statDeltaTimePause <= #TIME_PAUSE1_MAX))
                   THEN
                       #statChannelActive2 := true;
                       #statCountChannelPos := #CONST_CHANNEL_POS2; // go to next pos 2
                   END_IF;

                   IF ((#statDeltaTimePause >= #TIME_PAUSE2_MIN)
                       AND (#statDeltaTimePause <= #TIME_PAUSE2_MAX))
                   THEN
                       #statChannelActive2 := false;
                       #statChannelActive3 := true;
                       #statCountChannelPos := #CONST_CHANNEL_POS2; // go to next Pos 2
                   END_IF;

                   IF ((#statDeltaTimePause >= #TIME_PAUSE3_MIN)
                       AND (#statDeltaTimePause <= #TIME_PAUSE3_MAX))
                   THEN
                       #statChannelActive2 := false;
                       #statChannelActive3 := false;
                       #statChannelActive4 := true;
                       #statCountChannelPos := #CONST_INT_0;
                   END_IF;

               ELSIF (#statCountChannelPos = #CONST_CHANNEL_POS2)
               THEN
                   #statCurrentPos3 := #statCountChannelPos;
                   #statTimeImpulseSave3 := #statDeltaTimeImpulse;
                   #statTimePauseSave3 := #statDeltaTimePause;
                   #statTimeToImpulse := #statTimeToImpulse + #statDeltaTimeImpulse + #statDeltaTimePause;

                   IF ((#statDeltaTimePause >= #TIME_PAUSE1_MIN)
                       AND (#statDeltaTimePause <= #TIME_PAUSE1_MAX))
                   THEN
                       #statChannelActive3 := true;
                       #statCountChannelPos := #CONST_CHANNEL_POS3; // go to next pos 3
                   END_IF;

                   IF ((#statDeltaTimePause >= #TIME_PAUSE2_MIN)
                       AND (#statDeltaTimePause <= #TIME_PAUSE2_MAX))
                   THEN
                       #statChannelActive3 := false;
                       #statChannelActive4 := true;
                       #statCountChannelPos := #CONST_INT_0;
                   END_IF;

               ELSIF (#statCountChannelPos = #CONST_CHANNEL_POS3)
               THEN
                   #statCurrentPos4 := #statCountChannelPos;
                   #statTimeImpulseSave4 := #statDeltaTimeImpulse;
                   #statTimePauseSave4 := #statDeltaTimePause;
                   #statTimeToImpulse := #statTimeToImpulse + #statDeltaTimeImpulse + #statDeltaTimePause;

                   IF ((#statDeltaTimePause >= #TIME_PAUSE1_MIN)
                       AND (#statDeltaTimePause <= #TIME_PAUSE1_MAX))
                   THEN
                       #statChannelActive4 := true;
                   END_IF;
                   #statCountChannelPos := #CONST_INT_0; // go to pos 0
               END_IF;
           END_IF;

       #STATE_ERROR:
           #Error := true;
           #Busy := false;
           #Done := false;
           #statSysTimerStart := false;
           #statWatchDogTimerRisingStart := false;
           #statWatchDogTimerFallingStart := false;
           #Status := #statStatus;
           #statStatus := #CONST_WORD_0;
           #statIndex := #STATE_IDLE;
       ELSE
           #statIndex := #STATE_IDLE;
   END_CASE;

   #instWatchDogTimerRising(IN := #statWatchDogTimerRisingStart,
                      PT := #CONST_WATCHDOG_TIMER,
                      Q=>#statWatchDogTimerRisingStop,
                      ET=>#statWatchDogTimerRisingRun);

   #instWatchDogTimerFalling(IN:=#statWatchDogTimerFallingStart,
                             PT:=#CONST_WATCHDOG_TIMER,
                             Q=>#statWatchDogTimerFallingStop,
                             ET=>#statWatchDogTimerFallingRun);


   #instSysTimer(IN:=#statSysTimerStart,
                 PT:=#CONST_CYCLETIME_TIMER,
                 Q=>#statSysTimerStop,
                 ET=>#statSysTimerRun);

